DATA_BLOCK "DB619_State_MPart"   // DB619
TITLE = Status of maschine units and foaming cycle
{ S7_Optimized_Access := 'FALSE' }
VERSION : 0.1
   VAR
      ReadDeviceNo : Int := 1;
      ActualDeviceNo : Int := 0;
      CopyDeviceNO : Int := 0;
      Read : Bool := FALSE;
      Write : Bool := FALSE;
      Copy : Bool := FALSE;
      Operationmode : Array[0..2] of "UDT011_Operationmode";   // State operation mode machine
      Recirculation : Array[0..2] of "UDT012_Recirculation";   // State recirculation machine
      SWU : Array[0..2] of "UDT041_SWU_State";   // State selction switch over unit
      Mixinghead : Array[0..2] of "UDT042_MH_Select";   // State selection mixinghaead
      Cycle : Array[0..2] of "UDT091_PouringCycleState";   // State foaming cycle machine
      CylinderManager : Array[0..2] of "UDT061_Cylinder_Manager";   // State cylinder manager machine
      ToolMa : Array[0..2] of "UDT935_StatusShotSequenc";   // State of shot sequence machine
      ShotMa : Array[0..2] of Struct   // Shot values of machine 1 - 2
         Tool : "UDT926_ShotSet";
         ShotData : "UDT937_ShotData";
      END_STRUCT;
      PressureMHConnection : Array[0..8] of Real;   // Set values pressure at the connector of the mixinghead during a shot
      Machine : Array[0..2] of "UDT10_Machine";   // State of machine
      ActPressureMa : Array[0..2] of Struct   // Actual pressure at the MH-Connections of all 4 machines
         MH_Con : Array[1..8] of Real;   // values of the single connections
      END_STRUCT;
      ActMHPressureMa : Array[0..2] of Struct   // Actual pressure of the components involved at shot for each machine
         Comp : Array[1..12] of Real;   // single component value
      END_STRUCT;
      ActTemperatureMa : Array[0..2] of Struct   // Actual temperature at the MH-Connections of all 4 machines
         MH_Con : Array[1..8] of Real;   // values of the single connections
      END_STRUCT;
      ActMHTemperatureMa : Array[0..2] of Struct   // Actual temperature of the components involved at shot
         Comp : Array[1..12] of Real;   // single component value
      END_STRUCT;
      MH_at_Machine : Array[0..2] of "UDT001_DWord_1_32";   // Which mixinghead works at machine, Bit 0-31 corresponds to Mixinghead 1-32
      ActMixinghead : Array[0..8] of Int;
      BufferShotResultSignal : "UDT915_BuffResultSignal";   // State buffer shot results
      ActMHComponent : Array[0..2] of Struct
         No : Byte;
         OP_Manual : Bool;   // Opertaion mode manual at the mixinghead selected
         OP_Automatic : Bool;   // Opertaion mode automatic at the mixinghead selected
         OP_Service : Bool;   // Opertaion mode service (without foam) at the mixinghead selected
         Spare_4 : Bool;
         Spare_5 : Bool;
         Spare_6 : Bool;
         Spare_7 : Bool;
         Spare_8 : Bool;
         colour : Array[1..6] of Byte;
         "Name" : Array[1..6] of String[20];
      END_STRUCT;
      ActMHInerting : Array[0..2] of "UDT126_Inerting_ActValues_Ma";
      LP_Circ_Mixhead : Array[0..2] of "UDT014_LP_Circulation_MH";
   END_VAR
BEGIN
   Operationmode[0].valid := FALSE;
   Operationmode[0].Manual := FALSE;
   Operationmode[0].Auto := FALSE;
   Operationmode[0].Cylinderservice := FALSE;
   Operationmode[0].Test := FALSE;
   Operationmode[0].Operation := FALSE;
   Operationmode[0].Lamptest := FALSE;
   Operationmode[0].Controllvoltage := FALSE;
   Operationmode[0].Edge_OM_Change := FALSE;
   Operationmode[0].Active := FALSE;
   Operationmode[0].SwitchManual := FALSE;
   Operationmode[0].SwitchAutomatic := FALSE;
   Operationmode[0].SwitchOperation := FALSE;
   Operationmode[0].SwitchWeekEnd := FALSE;
   Operationmode[0].SwitchLamptest := FALSE;
   Operationmode[0].Spare16 := FALSE;
   Operationmode[1].valid := FALSE;
   Operationmode[1].Manual := FALSE;
   Operationmode[1].Auto := FALSE;
   Operationmode[1].Cylinderservice := FALSE;
   Operationmode[1].Test := FALSE;
   Operationmode[1].Operation := FALSE;
   Operationmode[1].Lamptest := FALSE;
   Operationmode[1].Controllvoltage := FALSE;
   Operationmode[1].Edge_OM_Change := FALSE;
   Operationmode[1].Active := FALSE;
   Operationmode[1].SwitchManual := FALSE;
   Operationmode[1].SwitchAutomatic := FALSE;
   Operationmode[1].SwitchOperation := FALSE;
   Operationmode[1].SwitchWeekEnd := FALSE;
   Operationmode[1].SwitchLamptest := FALSE;
   Operationmode[1].Spare16 := FALSE;
   Operationmode[2].valid := FALSE;
   Operationmode[2].Manual := FALSE;
   Operationmode[2].Auto := FALSE;
   Operationmode[2].Cylinderservice := FALSE;
   Operationmode[2].Test := FALSE;
   Operationmode[2].Operation := FALSE;
   Operationmode[2].Lamptest := FALSE;
   Operationmode[2].Controllvoltage := FALSE;
   Operationmode[2].Edge_OM_Change := FALSE;
   Operationmode[2].Active := FALSE;
   Operationmode[2].SwitchManual := FALSE;
   Operationmode[2].SwitchAutomatic := FALSE;
   Operationmode[2].SwitchOperation := FALSE;
   Operationmode[2].SwitchWeekEnd := FALSE;
   Operationmode[2].SwitchLamptest := FALSE;
   Operationmode[2].Spare16 := FALSE;
   Recirculation[0].Intervall := FALSE;
   Recirculation[0].Parallel := FALSE;
   Recirculation[0].Lowpressure := FALSE;
   Recirculation[0].Reduced := FALSE;
   Recirculation[0].Highpressure := FALSE;
   Recirculation[0].Tolerance_OK := FALSE;
   Recirculation[0].Weekendswitching := FALSE;
   Recirculation[0].Pausetime := FALSE;
   Recirculation[0].Break_KK := FALSE;
   Recirculation[0].HP_is_active := FALSE;
   Recirculation[0].Is_selected := FALSE;
   Recirculation[0].RequestPausePos := FALSE;
   Recirculation[0].cycle_runs := FALSE;
   Recirculation[0].Is_active := FALSE;
   Recirculation[0].Lowpressure_Exist := FALSE;
   Recirculation[0].Spare_1_7 := FALSE;
   Recirculation[0].Switch_Intervall := FALSE;
   Recirculation[0].Switch_Parallel := FALSE;
   Recirculation[0].Switch_Lowpressure := FALSE;
   Recirculation[0].Switch_Reduced := FALSE;
   Recirculation[0].Intervall_Reduced := FALSE;
   Recirculation[0].Intervall_Lowpressure := FALSE;
   Recirculation[0].Intervall_Reduced_Pause := FALSE;
   Recirculation[0].Intervall_Lowpressure_Pause := FALSE;
   Recirculation[0].Spare_3_0 := FALSE;
   Recirculation[0].Spare_3_1 := FALSE;
   Recirculation[0].Spare_3_2 := FALSE;
   Recirculation[0].Spare_3_3 := FALSE;
   Recirculation[0].Spare_3_4 := FALSE;
   Recirculation[0].Spare_3_5 := FALSE;
   Recirculation[0].Spare_3_6 := FALSE;
   Recirculation[0].Spare_3_7 := FALSE;
   Recirculation[0].State_Intervall := 0;
   Recirculation[0].State_Lowpressure := 0;
   Recirculation[0].State_Reduced := 0;
   Recirculation[0].Indicator_HP."25" := FALSE;
   Recirculation[0].Indicator_HP."26" := FALSE;
   Recirculation[0].Indicator_HP."27" := FALSE;
   Recirculation[0].Indicator_HP."28" := FALSE;
   Recirculation[0].Indicator_HP."29" := FALSE;
   Recirculation[0].Indicator_HP."30" := FALSE;
   Recirculation[0].Indicator_HP."31" := FALSE;
   Recirculation[0].Indicator_HP."32" := FALSE;
   Recirculation[0].Indicator_HP."17" := FALSE;
   Recirculation[0].Indicator_HP."18" := FALSE;
   Recirculation[0].Indicator_HP."19" := FALSE;
   Recirculation[0].Indicator_HP."20" := FALSE;
   Recirculation[0].Indicator_HP."21" := FALSE;
   Recirculation[0].Indicator_HP."22" := FALSE;
   Recirculation[0].Indicator_HP."23" := FALSE;
   Recirculation[0].Indicator_HP."24" := FALSE;
   Recirculation[0].Indicator_HP."09" := FALSE;
   Recirculation[0].Indicator_HP."10" := FALSE;
   Recirculation[0].Indicator_HP."11" := FALSE;
   Recirculation[0].Indicator_HP."12" := FALSE;
   Recirculation[0].Indicator_HP."13" := FALSE;
   Recirculation[0].Indicator_HP."14" := FALSE;
   Recirculation[0].Indicator_HP."15" := FALSE;
   Recirculation[0].Indicator_HP."16" := FALSE;
   Recirculation[0].Indicator_HP."01" := FALSE;
   Recirculation[0].Indicator_HP."02" := FALSE;
   Recirculation[0].Indicator_HP."03" := FALSE;
   Recirculation[0].Indicator_HP."04" := FALSE;
   Recirculation[0].Indicator_HP."05" := FALSE;
   Recirculation[0].Indicator_HP."06" := FALSE;
   Recirculation[0].Indicator_HP."07" := FALSE;
   Recirculation[0].Indicator_HP."08" := FALSE;
   Recirculation[0].Status_RC_HP := 0;
   Recirculation[0].Button_HP."25" := FALSE;
   Recirculation[0].Button_HP."26" := FALSE;
   Recirculation[0].Button_HP."27" := FALSE;
   Recirculation[0].Button_HP."28" := FALSE;
   Recirculation[0].Button_HP."29" := FALSE;
   Recirculation[0].Button_HP."30" := FALSE;
   Recirculation[0].Button_HP."31" := FALSE;
   Recirculation[0].Button_HP."32" := FALSE;
   Recirculation[0].Button_HP."17" := FALSE;
   Recirculation[0].Button_HP."18" := FALSE;
   Recirculation[0].Button_HP."19" := FALSE;
   Recirculation[0].Button_HP."20" := FALSE;
   Recirculation[0].Button_HP."21" := FALSE;
   Recirculation[0].Button_HP."22" := FALSE;
   Recirculation[0].Button_HP."23" := FALSE;
   Recirculation[0].Button_HP."24" := FALSE;
   Recirculation[0].Button_HP."09" := FALSE;
   Recirculation[0].Button_HP."10" := FALSE;
   Recirculation[0].Button_HP."11" := FALSE;
   Recirculation[0].Button_HP."12" := FALSE;
   Recirculation[0].Button_HP."13" := FALSE;
   Recirculation[0].Button_HP."14" := FALSE;
   Recirculation[0].Button_HP."15" := FALSE;
   Recirculation[0].Button_HP."16" := FALSE;
   Recirculation[0].Button_HP."01" := FALSE;
   Recirculation[0].Button_HP."02" := FALSE;
   Recirculation[0].Button_HP."03" := FALSE;
   Recirculation[0].Button_HP."04" := FALSE;
   Recirculation[0].Button_HP."05" := FALSE;
   Recirculation[0].Button_HP."06" := FALSE;
   Recirculation[0].Button_HP."07" := FALSE;
   Recirculation[0].Button_HP."08" := FALSE;
   Recirculation[0].Lamp_HP."25" := FALSE;
   Recirculation[0].Lamp_HP."26" := FALSE;
   Recirculation[0].Lamp_HP."27" := FALSE;
   Recirculation[0].Lamp_HP."28" := FALSE;
   Recirculation[0].Lamp_HP."29" := FALSE;
   Recirculation[0].Lamp_HP."30" := FALSE;
   Recirculation[0].Lamp_HP."31" := FALSE;
   Recirculation[0].Lamp_HP."32" := FALSE;
   Recirculation[0].Lamp_HP."17" := FALSE;
   Recirculation[0].Lamp_HP."18" := FALSE;
   Recirculation[0].Lamp_HP."19" := FALSE;
   Recirculation[0].Lamp_HP."20" := FALSE;
   Recirculation[0].Lamp_HP."21" := FALSE;
   Recirculation[0].Lamp_HP."22" := FALSE;
   Recirculation[0].Lamp_HP."23" := FALSE;
   Recirculation[0].Lamp_HP."24" := FALSE;
   Recirculation[0].Lamp_HP."09" := FALSE;
   Recirculation[0].Lamp_HP."10" := FALSE;
   Recirculation[0].Lamp_HP."11" := FALSE;
   Recirculation[0].Lamp_HP."12" := FALSE;
   Recirculation[0].Lamp_HP."13" := FALSE;
   Recirculation[0].Lamp_HP."14" := FALSE;
   Recirculation[0].Lamp_HP."15" := FALSE;
   Recirculation[0].Lamp_HP."16" := FALSE;
   Recirculation[0].Lamp_HP."01" := FALSE;
   Recirculation[0].Lamp_HP."02" := FALSE;
   Recirculation[0].Lamp_HP."03" := FALSE;
   Recirculation[0].Lamp_HP."04" := FALSE;
   Recirculation[0].Lamp_HP."05" := FALSE;
   Recirculation[0].Lamp_HP."06" := FALSE;
   Recirculation[0].Lamp_HP."07" := FALSE;
   Recirculation[0].Lamp_HP."08" := FALSE;
   Recirculation[0].SWU_RC_HP := 16#0000_0000;
   Recirculation[1].Intervall := FALSE;
   Recirculation[1].Parallel := FALSE;
   Recirculation[1].Lowpressure := FALSE;
   Recirculation[1].Reduced := FALSE;
   Recirculation[1].Highpressure := FALSE;
   Recirculation[1].Tolerance_OK := FALSE;
   Recirculation[1].Weekendswitching := FALSE;
   Recirculation[1].Pausetime := FALSE;
   Recirculation[1].Break_KK := FALSE;
   Recirculation[1].HP_is_active := FALSE;
   Recirculation[1].Is_selected := FALSE;
   Recirculation[1].RequestPausePos := FALSE;
   Recirculation[1].cycle_runs := FALSE;
   Recirculation[1].Is_active := FALSE;
   Recirculation[1].Lowpressure_Exist := FALSE;
   Recirculation[1].Spare_1_7 := FALSE;
   Recirculation[1].Switch_Intervall := FALSE;
   Recirculation[1].Switch_Parallel := FALSE;
   Recirculation[1].Switch_Lowpressure := FALSE;
   // 2234 more start values not shown
END_DATA_BLOCK

DATA_BLOCK "DB700_Machine"   // DB700
TITLE = Parameter PU machine
{ S7_Optimized_Access := 'FALSE' }
VERSION : 0.1
   VAR
      ReadWriteDeviceNo : Int := 1;
      CopyDeviceNO : Int := 0;
      Read : Bool := FALSE;
      Write : Bool := FALSE;
      Copy : Bool := FALSE;
      Machine : Array[0..2] of "UDT700_Machine";
   END_VAR
BEGIN
   Machine[1].Int_Runtime_Manual := S5T#30S;
   Machine[1].Int_Pausetime_Manual := S5T#30S;
   Machine[1].Int_Runtime_Auto := S5T#10S;
   Machine[1].Int_Pausetime_Auto := S5T#10S;
   Machine[1].SWU_Intervalltime := S5T#30S;
   Machine[1].HP_time_after_shot := S5T#10S;
   Machine[1].LP_Valve_switchOFF_Delay := S5T#30S;
   Machine[1].PressureBuildUpTime := S5T#10S;
   Machine[1].StandByTime := S5T#3S;
   Machine[1].CtrlChangeTime1 := S5T#3S;
   Machine[1].Max_ShotTime := S5T#34S;
   Machine[1].Max_WaitTime := S5T#1M;
   Machine[0].Int_Runtime_Manual := S5T#30S;
   Machine[0].Int_Pausetime_Manual := S5T#30S;
   Machine[0].Int_Runtime_Auto := S5T#10S;
   Machine[0].Int_Pausetime_Auto := S5T#10S;
   Machine[0].StrokeCounter_KK := 0;
   Machine[0].SWU_Intervalltime := S5T#30S;
   Machine[0].HP_time_after_shot := S5T#10S;
   Machine[0].LP_Valve_switchOFF_Delay := S5T#30S;
   Machine[0].PressureBuildUpTime := S5T#10S;
   Machine[0].StandByTime := S5T#3S;
   Machine[0].CtrlChangeTime1 := S5T#3S;
   Machine[0].Max_ShotTime := S5T#34S;
   Machine[0].Max_WaitTime := S5T#1M;
   Machine[0].MH_at_Machine := 16#0000_0001;
   Machine[0].Comp_at_Machine := 16#0000;
   Machine[0].CompPiston_at_Machine := 16#0000;
   Machine[1].StrokeCounter_KK := 0;
   Machine[1].MH_at_Machine := 16#0000_0001;
   Machine[1].Comp_at_Machine := 16#0000;
   Machine[1].CompPiston_at_Machine := 16#0000;
   Machine[2].Int_Runtime_Manual := S5T#0MS;
   Machine[2].Int_Pausetime_Manual := S5T#0MS;
   Machine[2].Int_Runtime_Auto := S5T#0MS;
   Machine[2].Int_Pausetime_Auto := S5T#0MS;
   Machine[2].StrokeCounter_KK := 0;
   Machine[2].SWU_Intervalltime := S5T#0MS;
   Machine[2].HP_time_after_shot := S5T#0MS;
   Machine[2].LP_Valve_switchOFF_Delay := S5T#0MS;
   Machine[2].PressureBuildUpTime := S5T#0MS;
   Machine[2].StandByTime := S5T#0MS;
   Machine[2].CtrlChangeTime1 := S5T#0MS;
   Machine[2].Max_ShotTime := S5T#0MS;
   Machine[2].Max_WaitTime := S5T#0MS;
   Machine[2].MH_at_Machine := 16#0000_0000;
   Machine[2].Comp_at_Machine := 16#0000;
   Machine[2].CompPiston_at_Machine := 16#0000;
   Machine[0].Min_ShotTime := S5T#200MS;
   Machine[1].Min_ShotTime := S5T#200MS;
   Machine[2].Min_ShotTime := S5T#0MS;
   Machine[0].CtrlChangeTime2 := S5T#600MS;
   Machine[1].CtrlChangeTime2 := S5T#600MS;
   Machine[2].CtrlChangeTime2 := S5T#0MS;
END_DATA_BLOCK

DATA_BLOCK "DB751_auxiliaryDriveMetering"   // DB701
TITLE = Parameter of universal drive
{ S7_Optimized_Access := 'FALSE' }
VERSION : 0.1
   VAR
      ReadWriteDeviceNo : Int := 0;
      CopyDeviceNO : Int := 0;
      Read : Bool := FALSE;
      Write : Bool := FALSE;
      Copy : Bool := FALSE;
      FeedingPump : Array[0..12] of "UDT710_FeedingPump";   // Pump to feed the metering pump
      EdgeFilter : Array[0..12] of "UDT710_EdgeFilter";
      HeatConverter : Array[0..12] of "UDT734_HeatConverter";
      HeatexchangerHP : Array[0..12] of "UDT780_ParaPW_Controller";
      HeatexchangerLP : Array[0..12] of "UDT780_ParaPW_Controller";
      FeedingPumpControler : Array[0..12] of "UDT781_ParaPID_Ctrl";
   END_VAR
BEGIN
   FeedingPump[0].Config_Exist := FALSE;
   FeedingPump[0].Config_WithFC := FALSE;
   FeedingPump[0].Config_Without_PresControl := FALSE;
   FeedingPump[0].Config_With_PresControl := FALSE;
   FeedingPump[0].Config_Bypass := FALSE;
   FeedingPump[0].Config_Filling := FALSE;
   FeedingPump[0].Config_ManualSwitchON := FALSE;
   FeedingPump[0].Config_Spare8 := FALSE;
   FeedingPump[0].Config_Spare9 := FALSE;
   FeedingPump[0].Config_Spare10 := FALSE;
   FeedingPump[0].Config_Spare11 := FALSE;
   FeedingPump[0].Config_Spare12 := FALSE;
   FeedingPump[0].Config_Spare13 := FALSE;
   FeedingPump[0].Config_Spare14 := FALSE;
   FeedingPump[0].Config_Spare15 := FALSE;
   FeedingPump[0].Config_Spare16 := FALSE;
   FeedingPump[0].RunTime := S5T#10S;
   FeedingPump[0].PauseTime := S5T#30S;
   FeedingPump[0].MinTempRelease := 0;
   FeedingPump[1].Config_Exist := FALSE;
   FeedingPump[1].Config_WithFC := FALSE;
   FeedingPump[1].Config_Without_PresControl := FALSE;
   FeedingPump[1].Config_With_PresControl := FALSE;
   FeedingPump[1].Config_Bypass := FALSE;
   FeedingPump[1].Config_Filling := FALSE;
   FeedingPump[1].Config_ManualSwitchON := FALSE;
   FeedingPump[1].Config_Spare8 := FALSE;
   FeedingPump[1].Config_Spare9 := FALSE;
   FeedingPump[1].Config_Spare10 := FALSE;
   FeedingPump[1].Config_Spare11 := FALSE;
   FeedingPump[1].Config_Spare12 := FALSE;
   FeedingPump[1].Config_Spare13 := FALSE;
   FeedingPump[1].Config_Spare14 := FALSE;
   FeedingPump[1].Config_Spare15 := FALSE;
   FeedingPump[1].Config_Spare16 := FALSE;
   FeedingPump[1].RunTime := S5T#10S;
   FeedingPump[1].PauseTime := S5T#30S;
   FeedingPump[1].MinTempRelease := 0;
   FeedingPump[2].Config_Exist := FALSE;
   FeedingPump[2].Config_WithFC := FALSE;
   FeedingPump[2].Config_Without_PresControl := FALSE;
   FeedingPump[2].Config_With_PresControl := FALSE;
   FeedingPump[2].Config_Bypass := FALSE;
   FeedingPump[2].Config_Filling := FALSE;
   FeedingPump[2].Config_ManualSwitchON := FALSE;
   FeedingPump[2].Config_Spare8 := FALSE;
   FeedingPump[2].Config_Spare9 := FALSE;
   FeedingPump[2].Config_Spare10 := FALSE;
   FeedingPump[2].Config_Spare11 := FALSE;
   FeedingPump[2].Config_Spare12 := FALSE;
   FeedingPump[2].Config_Spare13 := FALSE;
   FeedingPump[2].Config_Spare14 := FALSE;
   FeedingPump[2].Config_Spare15 := FALSE;
   FeedingPump[2].Config_Spare16 := FALSE;
   FeedingPump[2].RunTime := S5T#1M;
   FeedingPump[2].PauseTime := S5T#0MS;
   FeedingPump[2].MinTempRelease := 0;
   FeedingPump[3].Config_Exist := FALSE;
   FeedingPump[3].Config_WithFC := FALSE;
   FeedingPump[3].Config_Without_PresControl := FALSE;
   FeedingPump[3].Config_With_PresControl := FALSE;
   FeedingPump[3].Config_Bypass := FALSE;
   FeedingPump[3].Config_Filling := FALSE;
   FeedingPump[3].Config_ManualSwitchON := FALSE;
   FeedingPump[3].Config_Spare8 := FALSE;
   FeedingPump[3].Config_Spare9 := FALSE;
   FeedingPump[3].Config_Spare10 := FALSE;
   FeedingPump[3].Config_Spare11 := FALSE;
   FeedingPump[3].Config_Spare12 := FALSE;
   FeedingPump[3].Config_Spare13 := FALSE;
   FeedingPump[3].Config_Spare14 := FALSE;
   FeedingPump[3].Config_Spare15 := FALSE;
   FeedingPump[3].Config_Spare16 := FALSE;
   FeedingPump[3].RunTime := S5T#0MS;
   FeedingPump[3].PauseTime := S5T#0MS;
   FeedingPump[3].MinTempRelease := 0;
   FeedingPump[4].Config_Exist := FALSE;
   FeedingPump[4].Config_WithFC := FALSE;
   FeedingPump[4].Config_Without_PresControl := FALSE;
   FeedingPump[4].Config_With_PresControl := FALSE;
   FeedingPump[4].Config_Bypass := FALSE;
   FeedingPump[4].Config_Filling := FALSE;
   FeedingPump[4].Config_ManualSwitchON := FALSE;
   FeedingPump[4].Config_Spare8 := FALSE;
   FeedingPump[4].Config_Spare9 := FALSE;
   FeedingPump[4].Config_Spare10 := FALSE;
   FeedingPump[4].Config_Spare11 := FALSE;
   FeedingPump[4].Config_Spare12 := FALSE;
   FeedingPump[4].Config_Spare13 := FALSE;
   FeedingPump[4].Config_Spare14 := FALSE;
   FeedingPump[4].Config_Spare15 := FALSE;
   FeedingPump[4].Config_Spare16 := FALSE;
   FeedingPump[4].RunTime := S5T#0MS;
   FeedingPump[4].PauseTime := S5T#0MS;
   FeedingPump[4].MinTempRelease := 0;
   FeedingPump[5].Config_Exist := FALSE;
   FeedingPump[5].Config_WithFC := FALSE;
   FeedingPump[5].Config_Without_PresControl := FALSE;
   FeedingPump[5].Config_With_PresControl := FALSE;
   FeedingPump[5].Config_Bypass := FALSE;
   FeedingPump[5].Config_Filling := FALSE;
   FeedingPump[5].Config_ManualSwitchON := FALSE;
   FeedingPump[5].Config_Spare8 := FALSE;
   FeedingPump[5].Config_Spare9 := FALSE;
   FeedingPump[5].Config_Spare10 := FALSE;
   FeedingPump[5].Config_Spare11 := FALSE;
   FeedingPump[5].Config_Spare12 := FALSE;
   FeedingPump[5].Config_Spare13 := FALSE;
   FeedingPump[5].Config_Spare14 := FALSE;
   FeedingPump[5].Config_Spare15 := FALSE;
   FeedingPump[5].Config_Spare16 := FALSE;
   FeedingPump[5].RunTime := S5T#0MS;
   FeedingPump[5].PauseTime := S5T#0MS;
   FeedingPump[5].MinTempRelease := 0;
   FeedingPump[6].Config_Exist := FALSE;
   FeedingPump[6].Config_WithFC := FALSE;
   FeedingPump[6].Config_Without_PresControl := FALSE;
   FeedingPump[6].Config_With_PresControl := FALSE;
   FeedingPump[6].Config_Bypass := FALSE;
   FeedingPump[6].Config_Filling := FALSE;
   FeedingPump[6].Config_ManualSwitchON := FALSE;
   FeedingPump[6].Config_Spare8 := FALSE;
   FeedingPump[6].Config_Spare9 := FALSE;
   FeedingPump[6].Config_Spare10 := FALSE;
   FeedingPump[6].Config_Spare11 := FALSE;
   FeedingPump[6].Config_Spare12 := FALSE;
   FeedingPump[6].Config_Spare13 := FALSE;
   FeedingPump[6].Config_Spare14 := FALSE;
   FeedingPump[6].Config_Spare15 := FALSE;
   FeedingPump[6].Config_Spare16 := FALSE;
   FeedingPump[6].RunTime := S5T#0MS;
   FeedingPump[6].PauseTime := S5T#0MS;
   FeedingPump[6].MinTempRelease := 0;
   FeedingPump[7].Config_Exist := FALSE;
   FeedingPump[7].Config_WithFC := FALSE;
   FeedingPump[7].Config_Without_PresControl := FALSE;
   FeedingPump[7].Config_With_PresControl := FALSE;
   FeedingPump[7].Config_Bypass := FALSE;
   FeedingPump[7].Config_Filling := FALSE;
   FeedingPump[7].Config_ManualSwitchON := FALSE;
   FeedingPump[7].Config_Spare8 := FALSE;
   FeedingPump[7].Config_Spare9 := FALSE;
   FeedingPump[7].Config_Spare10 := FALSE;
   FeedingPump[7].Config_Spare11 := FALSE;
   FeedingPump[7].Config_Spare12 := FALSE;
   FeedingPump[7].Config_Spare13 := FALSE;
   FeedingPump[7].Config_Spare14 := FALSE;
   FeedingPump[7].Config_Spare15 := FALSE;
   FeedingPump[7].Config_Spare16 := FALSE;
   FeedingPump[7].RunTime := S5T#0MS;
   FeedingPump[7].PauseTime := S5T#0MS;
   FeedingPump[7].MinTempRelease := 0;
   FeedingPump[8].Config_Exist := FALSE;
   FeedingPump[8].Config_WithFC := FALSE;
   FeedingPump[8].Config_Without_PresControl := FALSE;
   FeedingPump[8].Config_With_PresControl := FALSE;
   FeedingPump[8].Config_Bypass := FALSE;
   FeedingPump[8].Config_Filling := FALSE;
   FeedingPump[8].Config_ManualSwitchON := FALSE;
   FeedingPump[8].Config_Spare8 := FALSE;
   FeedingPump[8].Config_Spare9 := FALSE;
   FeedingPump[8].Config_Spare10 := FALSE;
   FeedingPump[8].Config_Spare11 := FALSE;
   FeedingPump[8].Config_Spare12 := FALSE;
   FeedingPump[8].Config_Spare13 := FALSE;
   FeedingPump[8].Config_Spare14 := FALSE;
   FeedingPump[8].Config_Spare15 := FALSE;
   FeedingPump[8].Config_Spare16 := FALSE;
   FeedingPump[8].RunTime := S5T#0MS;
   FeedingPump[8].PauseTime := S5T#0MS;
   FeedingPump[8].MinTempRelease := 0;
   FeedingPump[9].Config_Exist := FALSE;
   FeedingPump[9].Config_WithFC := FALSE;
   FeedingPump[9].Config_Without_PresControl := FALSE;
   FeedingPump[9].Config_With_PresControl := FALSE;
   FeedingPump[9].Config_Bypass := FALSE;
   FeedingPump[9].Config_Filling := FALSE;
   FeedingPump[9].Config_ManualSwitchON := FALSE;
   FeedingPump[9].Config_Spare8 := FALSE;
   FeedingPump[9].Config_Spare9 := FALSE;
   FeedingPump[9].Config_Spare10 := FALSE;
   FeedingPump[9].Config_Spare11 := FALSE;
   FeedingPump[9].Config_Spare12 := FALSE;
   FeedingPump[9].Config_Spare13 := FALSE;
   FeedingPump[9].Config_Spare14 := FALSE;
   FeedingPump[9].Config_Spare15 := FALSE;
   FeedingPump[9].Config_Spare16 := FALSE;
   FeedingPump[9].RunTime := S5T#0MS;
   FeedingPump[9].PauseTime := S5T#0MS;
   FeedingPump[9].MinTempRelease := 0;
   FeedingPump[10].Config_Exist := FALSE;
   FeedingPump[10].Config_WithFC := FALSE;
   FeedingPump[10].Config_Without_PresControl := FALSE;
   FeedingPump[10].Config_With_PresControl := FALSE;
   FeedingPump[10].Config_Bypass := FALSE;
   FeedingPump[10].Config_Filling := FALSE;
   FeedingPump[10].Config_ManualSwitchON := FALSE;
   FeedingPump[10].Config_Spare8 := FALSE;
   FeedingPump[10].Config_Spare9 := FALSE;
   FeedingPump[10].Config_Spare10 := FALSE;
   // 398 more start values not shown
END_DATA_BLOCK

DATA_BLOCK "DB702_Tank_Value"   // DB702
TITLE = Parameter tank filling, material
{ S7_Optimized_Access := 'FALSE' }
NAME : Tank
VERSION : 0.1
   VAR
      ReadWriteDeviceNo : Int := 0;
      CopyDeviceNO : Int := 0;
      Read : Bool := FALSE;
      Write : Bool := FALSE;
      Copy : Bool := FALSE;
      Tank : Array[0..12] of "UDT702_Tank";
      AgitatorBarell : Array[0..12] of "UDT710_Agitator";
      Pt2_Controller : Array[0..12] of "UDT703_TemperingControl";
      Pt2_ControllerBarell : Array[0..12] of "UDT703_TemperingControl";
      CirculationPump : Array[0..12] of "UDT701_auxiliaryDrive";
   END_VAR
BEGIN
   Tank[1].Existing := TRUE;
   Tank[0]."Name" := 'Poly';
   Tank[0].FillingTimeControl := S5T#1M_40S;
   Tank[0].NoShotFilling := 0;
   Tank[0].TimeToStartFilling := S5T#0MS;
   Tank[0].PreAgitatingTime := S5T#0MS;
   Tank[0].Density := 1055;
   Tank[0].Existing := TRUE;
   Tank[0].DrainTank := FALSE;
   Tank[0].With_Level := TRUE;
   Tank[0].With_Level_Monitoring := FALSE;
   Tank[0].WIth_Loading := FALSE;
   Tank[0].With_Heating := TRUE;
   Tank[0].With_Vacuum := FALSE;
   Tank[0].With_Nucleation := FALSE;
   Tank[0].With_Heater_Returnline := FALSE;
   Tank[0].With_Drain := FALSE;
   Tank[0].With_ContainerStation := FALSE;
   Tank[0].With_BarelStationAgitator := FALSE;
   Tank[0].With_Level_3Liq := FALSE;
   Tank[0].With_Level_4Liq := FALSE;
   Tank[0].With_Level_Probe := TRUE;
   Tank[0].With_Level_SMin := FALSE;
   Tank[0].With_Level_SMax := TRUE;
   Tank[0].With_Triptray := FALSE;
   Tank[0].With_Level_Spare7 := FALSE;
   Tank[0].With_Level_Spare8 := FALSE;
   Tank[0].With_Filling := TRUE;
   Tank[0].With_Filling_Valve := TRUE;
   Tank[0].With_Filling_2Valve := FALSE;
   Tank[0].With_Filling_ShutDown := FALSE;
   Tank[0].With_Filling_Switch := FALSE;
   Tank[0].With_Filling_Pump := FALSE;
   Tank[0].With_Filling_DryRun := FALSE;
   Tank[0].With_Filling_Pentane := FALSE;
   Tank[0].With_Tempering := TRUE;
   Tank[0].With_Tempering_TempGeraet := FALSE;
   Tank[0].With_Tempering_VKaltwasser := TRUE;
   Tank[0].With_Tempering_Heizung := TRUE;
   Tank[0].With_Tempering_WTRL := TRUE;
   Tank[0].With_Tempering_WTmitFischer := FALSE;
   Tank[0].With_Tempering_WTBypass := FALSE;
   Tank[0].With_Tempering_WTVL := FALSE;
   Tank[0].With_BarelStation := FALSE;
   Tank[0].With_BarelStation_Zirkulation := FALSE;
   Tank[0].With_BarelStation_PnPump := TRUE;
   Tank[0].With_BarelStation_ElPump := FALSE;
   Tank[0].With_BarelStation_PnRW := FALSE;
   Tank[0].With_BarelStation_ElRW := FALSE;
   Tank[0].With_BarelStation_Heating := FALSE;
   Tank[0].With_BarelStation_HeatingBottom := FALSE;
   Tank[0].With_Agitator := TRUE;
   Tank[0].With_Agitator_Converter := FALSE;
   Tank[0].With_Agitator_SetValue := FALSE;
   Tank[0].With_Agitator_6SetValue := FALSE;
   Tank[0].With_Agitator_Spare5 := FALSE;
   Tank[0].With_Agitator_Spare6 := FALSE;
   Tank[0].With_Agitator_Spare7 := FALSE;
   Tank[0].With_Agitator_Spare8 := FALSE;
   Tank[0].Agitator.Config_bit_Converter := FALSE;
   Tank[0].Agitator.Config_bit_Converter_SW := FALSE;
   Tank[0].Agitator.Config_bit_Heating_ON := TRUE;
   Tank[0].Agitator.config_bit_Heating_Int := TRUE;
   Tank[0].Agitator.Config_bit_Cooling_ON := TRUE;
   Tank[0].Agitator.Config_bit_Cooling_Int := FALSE;
   Tank[0].Agitator.Config_bit_Filling_ON := TRUE;
   Tank[0].Agitator.Config_bit_Filling_Int := TRUE;
   Tank[0].Agitator.Config_bit_Charging_ON := FALSE;
   Tank[0].Agitator.Config_bit_Charging_Int := FALSE;
   Tank[0].Agitator.RunTime := S5T#10S;
   Tank[0].Agitator.PauseTime := S5T#20S;
   Tank[0].Agitator_BarelStation.Config_bit_Converter := FALSE;
   Tank[0].Agitator_BarelStation.Config_bit_Converter_SW := FALSE;
   Tank[0].Agitator_BarelStation.Config_bit_Heating_ON := FALSE;
   Tank[0].Agitator_BarelStation.config_bit_Heating_Int := FALSE;
   Tank[0].Agitator_BarelStation.Config_bit_Cooling_ON := FALSE;
   Tank[0].Agitator_BarelStation.Config_bit_Cooling_Int := FALSE;
   Tank[0].Agitator_BarelStation.Config_bit_Filling_ON := FALSE;
   Tank[0].Agitator_BarelStation.Config_bit_Filling_Int := FALSE;
   Tank[0].Agitator_BarelStation.Config_bit_Charging_ON := FALSE;
   Tank[0].Agitator_BarelStation.Config_bit_Charging_Int := FALSE;
   Tank[0].Agitator_BarelStation.RunTime := S5T#0MS;
   Tank[0].Agitator_BarelStation.PauseTime := S5T#0MS;
   Tank[1]."Name" := 'Poly';
   Tank[1].FillingTimeControl := S5T#1M_40S;
   Tank[1].NoShotFilling := 0;
   Tank[1].TimeToStartFilling := S5T#0MS;
   Tank[1].PreAgitatingTime := S5T#0MS;
   Tank[1].Density := 1055;
   Tank[1].DrainTank := FALSE;
   Tank[1].With_Level := TRUE;
   Tank[1].With_Level_Monitoring := FALSE;
   Tank[1].WIth_Loading := FALSE;
   Tank[1].With_Heating := TRUE;
   Tank[1].With_Vacuum := FALSE;
   Tank[1].With_Nucleation := FALSE;
   Tank[1].With_Heater_Returnline := FALSE;
   Tank[1].With_Drain := FALSE;
   Tank[1].With_ContainerStation := FALSE;
   Tank[1].With_BarelStationAgitator := FALSE;
   Tank[1].With_Level_3Liq := FALSE;
   Tank[1].With_Level_4Liq := FALSE;
   Tank[1].With_Level_Probe := TRUE;
   Tank[1].With_Level_SMin := FALSE;
   Tank[1].With_Level_SMax := TRUE;
   Tank[1].With_Triptray := FALSE;
   Tank[1].With_Level_Spare7 := FALSE;
   Tank[1].With_Level_Spare8 := FALSE;
   Tank[1].With_Filling := TRUE;
   Tank[1].With_Filling_Valve := TRUE;
   Tank[1].With_Filling_2Valve := FALSE;
   Tank[1].With_Filling_ShutDown := FALSE;
   Tank[1].With_Filling_Switch := FALSE;
   Tank[1].With_Filling_Pump := FALSE;
   Tank[1].With_Filling_DryRun := FALSE;
   Tank[1].With_Filling_Pentane := FALSE;
   Tank[1].With_Tempering := TRUE;
   Tank[1].With_Tempering_TempGeraet := FALSE;
   Tank[1].With_Tempering_VKaltwasser := TRUE;
   Tank[1].With_Tempering_Heizung := TRUE;
   Tank[1].With_Tempering_WTRL := TRUE;
   Tank[1].With_Tempering_WTmitFischer := FALSE;
   Tank[1].With_Tempering_WTBypass := FALSE;
   Tank[1].With_Tempering_WTVL := FALSE;
   Tank[1].With_BarelStation := FALSE;
   Tank[1].With_BarelStation_Zirkulation := FALSE;
   Tank[1].With_BarelStation_PnPump := TRUE;
   Tank[1].With_BarelStation_ElPump := FALSE;
   Tank[1].With_BarelStation_PnRW := FALSE;
   Tank[1].With_BarelStation_ElRW := FALSE;
   Tank[1].With_BarelStation_Heating := FALSE;
   Tank[1].With_BarelStation_HeatingBottom := FALSE;
   Tank[1].With_Agitator := TRUE;
   Tank[1].With_Agitator_Converter := FALSE;
   Tank[1].With_Agitator_SetValue := FALSE;
   Tank[1].With_Agitator_6SetValue := FALSE;
   Tank[1].With_Agitator_Spare5 := FALSE;
   Tank[1].With_Agitator_Spare6 := FALSE;
   Tank[1].With_Agitator_Spare7 := FALSE;
   Tank[1].With_Agitator_Spare8 := FALSE;
   Tank[1].Agitator.Config_bit_Converter := FALSE;
   Tank[1].Agitator.Config_bit_Converter_SW := FALSE;
   Tank[1].Agitator.Config_bit_Heating_ON := TRUE;
   Tank[1].Agitator.config_bit_Heating_Int := TRUE;
   Tank[1].Agitator.Config_bit_Cooling_ON := TRUE;
   Tank[1].Agitator.Config_bit_Cooling_Int := FALSE;
   Tank[1].Agitator.Config_bit_Filling_ON := TRUE;
   Tank[1].Agitator.Config_bit_Filling_Int := TRUE;
   Tank[1].Agitator.Config_bit_Charging_ON := FALSE;
   Tank[1].Agitator.Config_bit_Charging_Int := FALSE;
   Tank[1].Agitator.RunTime := S5T#10S;
   Tank[1].Agitator.PauseTime := S5T#20S;
   Tank[1].Agitator_BarelStation.Config_bit_Converter := FALSE;
   Tank[1].Agitator_BarelStation.Config_bit_Converter_SW := FALSE;
   Tank[1].Agitator_BarelStation.Config_bit_Heating_ON := FALSE;
   Tank[1].Agitator_BarelStation.config_bit_Heating_Int := FALSE;
   Tank[1].Agitator_BarelStation.Config_bit_Cooling_ON := FALSE;
   Tank[1].Agitator_BarelStation.Config_bit_Cooling_Int := FALSE;
   Tank[1].Agitator_BarelStation.Config_bit_Filling_ON := FALSE;
   Tank[1].Agitator_BarelStation.Config_bit_Filling_Int := FALSE;
   Tank[1].Agitator_BarelStation.Config_bit_Charging_ON := FALSE;
   Tank[1].Agitator_BarelStation.Config_bit_Charging_Int := FALSE;
   Tank[1].Agitator_BarelStation.RunTime := S5T#0MS;
   Tank[1].Agitator_BarelStation.PauseTime := S5T#0MS;
   Tank[2]."Name" := 'Iso';
   Tank[2].FillingTimeControl := S5T#1M_40S;
   Tank[2].NoShotFilling := 0;
   Tank[2].TimeToStartFilling := S5T#0MS;
   Tank[2].PreAgitatingTime := S5T#0MS;
   Tank[2].Density := 1055;
   Tank[2].Existing := TRUE;
   Tank[2].DrainTank := FALSE;
   Tank[2].With_Level := TRUE;
   Tank[2].With_Level_Monitoring := FALSE;
   Tank[2].WIth_Loading := FALSE;
   Tank[2].With_Heating := TRUE;
   Tank[2].With_Vacuum := FALSE;
   Tank[2].With_Nucleation := FALSE;
   Tank[2].With_Heater_Returnline := FALSE;
   Tank[2].With_Drain := FALSE;
   Tank[2].With_ContainerStation := FALSE;
   Tank[2].With_BarelStationAgitator := FALSE;
   Tank[2].With_Level_3Liq := FALSE;
   Tank[2].With_Level_4Liq := FALSE;
   Tank[2].With_Level_Probe := TRUE;
   Tank[2].With_Level_SMin := FALSE;
   Tank[2].With_Level_SMax := TRUE;
   Tank[2].With_Triptray := FALSE;
   Tank[2].With_Level_Spare7 := FALSE;
   Tank[2].With_Level_Spare8 := FALSE;
   Tank[2].With_Filling := TRUE;
   Tank[2].With_Filling_Valve := TRUE;
   Tank[2].With_Filling_2Valve := FALSE;
   Tank[2].With_Filling_ShutDown := FALSE;
   Tank[2].With_Filling_Switch := FALSE;
   Tank[2].With_Filling_Pump := FALSE;
   Tank[2].With_Filling_DryRun := FALSE;
   Tank[2].With_Filling_Pentane := FALSE;
   Tank[2].With_Tempering := TRUE;
   Tank[2].With_Tempering_TempGeraet := FALSE;
   // 1360 more start values not shown
END_DATA_BLOCK

DATA_BLOCK "DB704_MH_Value"   // DB704
TITLE = Parameter mixinghead
{ S7_Optimized_Access := 'FALSE' }
VERSION : 0.1
   VAR
      ReadWriteDeviceNo : Int := 0;
      CopyDeviceNO : Int := 0;
      Read : Bool := FALSE;
      Write : Bool := FALSE;
      Copy : Bool := FALSE;
      Mixinghead : Array[0..16] of "UDT704_Mixinghead";
      MH_Inerting : Array[0..16] of "UDT125_Inerting_SetValues";
   END_VAR
BEGIN
   Mixinghead[0].AmountComponent := 16#02;
   Mixinghead[0].MachineNumber := 16#01;
   Mixinghead[0].pRrgNumberManual := 16#00;
   Mixinghead[0].MH_Active := TRUE;
   Mixinghead[0].WithCleaningPiston := TRUE;
   Mixinghead[0].WithNozzleControl := FALSE;
   Mixinghead[0].WithLPCirculation := TRUE;
   Mixinghead[0].WithInterface := FALSE;
   Mixinghead[0].WithInerting := FALSE;
   Mixinghead[0].WithHeating := FALSE;
   Mixinghead[0].WithMHVenting := FALSE;
   Mixinghead[0].NozzleLeakageTest := FALSE;
   Mixinghead[0].ShotBreak := FALSE;
   Mixinghead[0].Conf_IntWithRobot := FALSE;
   Mixinghead[0].Conf_IntWithMC := FALSE;
   Mixinghead[0].Conf_IntWithPlantInerface := FALSE;
   Mixinghead[0].Conf_IntWithCoupler := FALSE;
   Mixinghead[0].Conf_MHDigital := TRUE;
   Mixinghead[0].Conf_MHControled := FALSE;
   Mixinghead[0].Conf_MHFibre := FALSE;
   Mixinghead[0].Conf_MHSpray := FALSE;
   Mixinghead[0].Conf_MHSpecial := FALSE;
   Mixinghead[0].Openingtime := 0.0;
   Mixinghead[0].Closingtime := 0.0;
   Mixinghead[0].NozzelCirc := 16#00;
   Mixinghead[0].NozzelShot := 16#00;
   Mixinghead[0].NozzleRelease := 16#00;
   Mixinghead[0].NozzelForcen := 16#00;
   Mixinghead[0].DelayTimeNozzlesOff := S5T#5S;
   Mixinghead[0].Delay_UnLockMHafterShot := S5T#0MS;
   Mixinghead[0].RunTime_MHLock := S5T#0MS;
   Mixinghead[0].RunTime_MHUnLock := S5T#0MS;
   Mixinghead[0].Cleaning_Piston.Offset_CP := 0;
   Mixinghead[0].Cleaning_Piston.Length_DrainPipe := 0;
   Mixinghead[0].Cleaning_Piston.Diam_Piston := 0;
   Mixinghead[0].Cleaning_Piston.ChokeSlot_min := 0;
   Mixinghead[0].Cleaning_Piston.ChokeSlot_max := 0;
   Mixinghead[0].Cleaning_Piston.RestTimeBack := S5T#200MS;
   Mixinghead[0].Cleaning_Piston.RestTimeFront := S5T#5S;
   Mixinghead[0].Cleaning_Piston.RestTimeFrontManual := S5T#5S;
   Mixinghead[0].Cleaning_Piston.IntervalCounts := 0;
   Mixinghead[0].Cleaning_Piston.IntervalRestTimeBack := S5T#0MS;
   Mixinghead[0].Cleaning_Piston.IntervalRestTimeFront := S5T#0MS;
   Mixinghead[0].Cleaning_Piston.CP_after_PS := FALSE;
   Mixinghead[0].Cleaning_Piston.CP_withInterval := FALSE;
   Mixinghead[0].Cleaning_Piston.StepCleaningPiston := FALSE;
   Mixinghead[0].Cleaning_Piston.ContrCleaningPiston := FALSE;
   Mixinghead[0].Cleaning_Piston.Spare_19 := FALSE;
   Mixinghead[0].Cleaning_Piston.Spare_20 := FALSE;
   Mixinghead[0].Cleaning_Piston.Spare_21 := FALSE;
   Mixinghead[0].Cleaning_Piston.Spare_22 := FALSE;
   Mixinghead[0].Cleaning_Piston.Spare_23 := FALSE;
   Mixinghead[0].Cleaning_Piston.Spare_24 := FALSE;
   Mixinghead[0].Cleaning_Piston.Spare_25 := FALSE;
   Mixinghead[0].Cleaning_Piston.Spare_26 := FALSE;
   Mixinghead[0].Cleaning_Piston.Spare_27 := FALSE;
   Mixinghead[0].Cleaning_Piston.Spare_28 := FALSE;
   Mixinghead[0].Cleaning_Piston.Spare_29 := FALSE;
   Mixinghead[0].Cleaning_Piston.Spare_30 := FALSE;
   Mixinghead[0].Steering_Piston.T_monitoring_open := S5T#0MS;
   Mixinghead[0].Steering_Piston.T_monitoring_close := S5T#0MS;
   Mixinghead[0].Corrvalue := 0.022;
   Mixinghead[0].Leading_Comp_No := 0;
   Mixinghead[0].MH_Connection[1].Pump_No := 1;
   Mixinghead[0].MH_Connection[1].Flow_HP_Circ := 400.0;
   Mixinghead[0].MH_Connection[1].Flow_red_Circ := 200.0;
   Mixinghead[0].MH_Connection[1].Flow_LP_Circ := 140.0;
   Mixinghead[0].MH_Connection[1].Nozzel_delay_open := 0.0;
   Mixinghead[0].MH_Connection[1].Nozzel_delay_close := 0.0;
   Mixinghead[0].MH_Connection[1].FlowQPB := 100.0;
   Mixinghead[0].MH_Connection[1].PressureQPB := 0.0;
   Mixinghead[0].MH_Connection[1].HP_CircOverNozzle := FALSE;
   Mixinghead[0].MH_Connection[1].Red_CircOverNozzle := FALSE;
   Mixinghead[0].MH_Connection[1].LP_CircOverNozzle := FALSE;
   Mixinghead[0].MH_Connection[1].WithNozzle := TRUE;
   Mixinghead[0].MH_Connection[1].HP_2Point_Flow := FALSE;
   Mixinghead[0].MH_Connection[1].Red_2Point_Flow := FALSE;
   Mixinghead[0].MH_Connection[1].LP_2Point_Flow := FALSE;
   Mixinghead[0].MH_Connection[1].Exist := TRUE;
   Mixinghead[0].MH_Connection[1].Spare27 := 16#00;
   Mixinghead[0].MH_Connection[2].Pump_No := 2;
   Mixinghead[0].MH_Connection[2].Flow_HP_Circ := 175.0;
   Mixinghead[0].MH_Connection[2].Flow_red_Circ := 100.0;
   Mixinghead[0].MH_Connection[2].Flow_LP_Circ := 75.0;
   Mixinghead[0].MH_Connection[2].Nozzel_delay_open := 0.0;
   Mixinghead[0].MH_Connection[2].Nozzel_delay_close := 0.0;
   Mixinghead[0].MH_Connection[2].FlowQPB := 100.0;
   Mixinghead[0].MH_Connection[2].PressureQPB := 0.0;
   Mixinghead[0].MH_Connection[2].HP_CircOverNozzle := FALSE;
   Mixinghead[0].MH_Connection[2].Red_CircOverNozzle := FALSE;
   Mixinghead[0].MH_Connection[2].LP_CircOverNozzle := FALSE;
   Mixinghead[0].MH_Connection[2].WithNozzle := TRUE;
   Mixinghead[0].MH_Connection[2].HP_2Point_Flow := FALSE;
   Mixinghead[0].MH_Connection[2].Red_2Point_Flow := FALSE;
   Mixinghead[0].MH_Connection[2].LP_2Point_Flow := FALSE;
   Mixinghead[0].MH_Connection[2].Exist := TRUE;
   Mixinghead[0].MH_Connection[2].Spare27 := 16#00;
   Mixinghead[0].MH_Connection[3].Pump_No := 0;
   Mixinghead[0].MH_Connection[3].Flow_HP_Circ := 0.0;
   Mixinghead[0].MH_Connection[3].Flow_red_Circ := 0.0;
   Mixinghead[0].MH_Connection[3].Flow_LP_Circ := 0.0;
   Mixinghead[0].MH_Connection[3].Nozzel_delay_open := 0.0;
   Mixinghead[0].MH_Connection[3].Nozzel_delay_close := 0.0;
   Mixinghead[0].MH_Connection[3].FlowQPB := 0.0;
   Mixinghead[0].MH_Connection[3].PressureQPB := 0.0;
   Mixinghead[0].MH_Connection[3].HP_CircOverNozzle := FALSE;
   Mixinghead[0].MH_Connection[3].Red_CircOverNozzle := FALSE;
   Mixinghead[0].MH_Connection[3].LP_CircOverNozzle := FALSE;
   Mixinghead[0].MH_Connection[3].WithNozzle := FALSE;
   Mixinghead[0].MH_Connection[3].HP_2Point_Flow := FALSE;
   Mixinghead[0].MH_Connection[3].Red_2Point_Flow := FALSE;
   Mixinghead[0].MH_Connection[3].LP_2Point_Flow := FALSE;
   Mixinghead[0].MH_Connection[3].Exist := FALSE;
   Mixinghead[0].MH_Connection[3].Spare27 := 16#00;
   Mixinghead[0].MH_Connection[4].Pump_No := 0;
   Mixinghead[0].MH_Connection[4].Flow_HP_Circ := 0.0;
   Mixinghead[0].MH_Connection[4].Flow_red_Circ := 0.0;
   Mixinghead[0].MH_Connection[4].Flow_LP_Circ := 0.0;
   Mixinghead[0].MH_Connection[4].Nozzel_delay_open := 0.0;
   Mixinghead[0].MH_Connection[4].Nozzel_delay_close := 0.0;
   Mixinghead[0].MH_Connection[4].FlowQPB := 0.0;
   Mixinghead[0].MH_Connection[4].PressureQPB := 0.0;
   Mixinghead[0].MH_Connection[4].HP_CircOverNozzle := FALSE;
   Mixinghead[0].MH_Connection[4].Red_CircOverNozzle := FALSE;
   Mixinghead[0].MH_Connection[4].LP_CircOverNozzle := FALSE;
   Mixinghead[0].MH_Connection[4].WithNozzle := FALSE;
   Mixinghead[0].MH_Connection[4].HP_2Point_Flow := FALSE;
   Mixinghead[0].MH_Connection[4].Red_2Point_Flow := FALSE;
   Mixinghead[0].MH_Connection[4].LP_2Point_Flow := FALSE;
   Mixinghead[0].MH_Connection[4].Exist := FALSE;
   Mixinghead[0].MH_Connection[4].Spare27 := 16#00;
   Mixinghead[0].MH_Connection[5].Pump_No := 0;
   Mixinghead[0].MH_Connection[5].Flow_HP_Circ := 0.0;
   Mixinghead[0].MH_Connection[5].Flow_red_Circ := 0.0;
   Mixinghead[0].MH_Connection[5].Flow_LP_Circ := 0.0;
   Mixinghead[0].MH_Connection[5].Nozzel_delay_open := 0.0;
   Mixinghead[0].MH_Connection[5].Nozzel_delay_close := 0.0;
   Mixinghead[0].MH_Connection[5].FlowQPB := 0.0;
   Mixinghead[0].MH_Connection[5].PressureQPB := 0.0;
   Mixinghead[0].MH_Connection[5].HP_CircOverNozzle := FALSE;
   Mixinghead[0].MH_Connection[5].Red_CircOverNozzle := FALSE;
   Mixinghead[0].MH_Connection[5].LP_CircOverNozzle := FALSE;
   Mixinghead[0].MH_Connection[5].WithNozzle := FALSE;
   Mixinghead[0].MH_Connection[5].HP_2Point_Flow := FALSE;
   Mixinghead[0].MH_Connection[5].Red_2Point_Flow := FALSE;
   Mixinghead[0].MH_Connection[5].LP_2Point_Flow := FALSE;
   Mixinghead[0].MH_Connection[5].Exist := FALSE;
   Mixinghead[0].MH_Connection[5].Spare27 := 16#00;
   Mixinghead[0].MH_Connection[6].Pump_No := 0;
   Mixinghead[0].MH_Connection[6].Flow_HP_Circ := 0.0;
   Mixinghead[0].MH_Connection[6].Flow_red_Circ := 0.0;
   Mixinghead[0].MH_Connection[6].Flow_LP_Circ := 0.0;
   Mixinghead[0].MH_Connection[6].Nozzel_delay_open := 0.0;
   Mixinghead[0].MH_Connection[6].Nozzel_delay_close := 0.0;
   Mixinghead[0].MH_Connection[6].FlowQPB := 0.0;
   Mixinghead[0].MH_Connection[6].PressureQPB := 0.0;
   Mixinghead[0].MH_Connection[6].HP_CircOverNozzle := FALSE;
   Mixinghead[0].MH_Connection[6].Red_CircOverNozzle := FALSE;
   Mixinghead[0].MH_Connection[6].LP_CircOverNozzle := FALSE;
   Mixinghead[0].MH_Connection[6].WithNozzle := FALSE;
   Mixinghead[0].MH_Connection[6].HP_2Point_Flow := FALSE;
   Mixinghead[0].MH_Connection[6].Red_2Point_Flow := FALSE;
   Mixinghead[0].MH_Connection[6].LP_2Point_Flow := FALSE;
   Mixinghead[0].MH_Connection[6].Exist := FALSE;
   Mixinghead[0].MH_Connection[6].Spare27 := 16#00;
   Mixinghead[1].AmountComponent := 16#02;
   Mixinghead[1].MachineNumber := 16#01;
   Mixinghead[1].pRrgNumberManual := 16#00;
   Mixinghead[1].MH_Active := TRUE;
   Mixinghead[1].WithCleaningPiston := TRUE;
   Mixinghead[1].WithNozzleControl := FALSE;
   Mixinghead[1].WithLPCirculation := TRUE;
   Mixinghead[1].WithInterface := FALSE;
   Mixinghead[1].WithInerting := FALSE;
   Mixinghead[1].WithHeating := FALSE;
   Mixinghead[1].WithMHVenting := FALSE;
   Mixinghead[1].NozzleLeakageTest := FALSE;
   Mixinghead[1].ShotBreak := FALSE;
   Mixinghead[1].Conf_IntWithRobot := FALSE;
   Mixinghead[1].Conf_IntWithMC := FALSE;
   Mixinghead[1].Conf_IntWithPlantInerface := FALSE;
   Mixinghead[1].Conf_IntWithCoupler := FALSE;
   Mixinghead[1].Conf_MHDigital := TRUE;
   Mixinghead[1].Conf_MHControled := FALSE;
   Mixinghead[1].Conf_MHFibre := FALSE;
   Mixinghead[1].Conf_MHSpray := FALSE;
   Mixinghead[1].Conf_MHSpecial := FALSE;
   Mixinghead[1].Openingtime := 0.0;
   Mixinghead[1].Closingtime := 0.0;
   Mixinghead[1].NozzelCirc := 16#00;
   Mixinghead[1].NozzelShot := 16#00;
   Mixinghead[1].NozzleRelease := 16#00;
   Mixinghead[1].NozzelForcen := 16#00;
   Mixinghead[1].DelayTimeNozzlesOff := S5T#5S;
   Mixinghead[1].Delay_UnLockMHafterShot := S5T#0MS;
   Mixinghead[1].RunTime_MHLock := S5T#0MS;
   Mixinghead[1].RunTime_MHUnLock := S5T#0MS;
   Mixinghead[1].Cleaning_Piston.Offset_CP := 0;
   Mixinghead[1].Cleaning_Piston.Length_DrainPipe := 0;
   Mixinghead[1].Cleaning_Piston.Diam_Piston := 0;
   // 4152 more start values not shown
END_DATA_BLOCK

DATA_BLOCK "DB721_MH_Hydraulic"   // DB721
TITLE = Parameter mixing head hydraulic
{ S7_Optimized_Access := 'FALSE' }
NAME : Hydrauli